VAR_GLOBAL CONSTANT   // PLC tag table "Open Library"
   "Modes.Auto" : Int := 1;
   "Modes.Manual" : Int := 2;
   "Modes.Independent" : Int := 10;
   "Modes.Stop" : Int := 0;
   "HMI.Status.Stopped" : Int := 0;
   "HMI.Status.Estop" : Int := 1;
   "HMI.Status.Error" : Int := 2;
   "HMI.Status.ForwardWork" : Int := 3;
   "HMI.Status.ReverseHome" : Int := 4;
   "HMI.Status.OnForwardWork" : Int := 5;
   "HMI.Status.OnReverseHome" : Int := 6;
   "IoScaling.S7Analog.Default.iRawMax" : Int := 27648;
   "IoScaling.S7Analog.Default.iRawMin" : Int := 0;
   "IoScaling.S7Analog.Default.bSwapBytes" : Bool := false;
   "IoScaling.S7Analog.+-V/mA.iRawMax" : Int := 27648;
   "IoScaling.S7Analog.+-V/mA.iRawMin" : Int := -27648;
   "IoScaling.S7Analog.Types.Default" : Int := 0;
   "IoScaling.S7Analog.Pt100.iRawMax" : Int := 8500;
   "IoScaling.S7Analog.Pt100.iRawMin" : Int := -2000;
   "IoScaling.S7Analog.Pt100.Climate.iRawMax" : Int := 13000;
   "IoScaling.S7Analog.Pt100.Climate.iRawMin" : Int := -12000;
   "IoScaling.S7Analog.Ni100.iRawMax" : Int := 2500;
   "IoScaling.S7Analog.Ni100.iRawMin" : Int := -600;
   "IoScaling.S7Analog.Ni100.Climate.iRawMax" : Int := 25000;
   "IoScaling.S7Analog.Ni100.Climate.iRawMin" : Int := -6000;
   "IoScaling.S7Analog.Types.+-V/mA" : Int := 1;
   "IoScaling.S7Analog.Types.Pt100" : Int := 2;
   "IoScaling.S7Analog.Types.Pt100.Climate" : Int := 3;
   "IoScaling.S7Analog.Types.Ni100" : Int := 4;
   "IoScaling.S7Analog.Types.Ni100.Climate" : Int := 5;
   "IoScaling.S7Analog.Pt100.rScaledMax" : Real := 850.0;
   "IoScaling.S7Analog.Pt100.rScaledMin" : Real := -200.0;
   "IoScaling.S7Analog.Pt100.Climate.rScaledMax" : Real := 130.0;
   "IoScaling.S7Analog.Pt100.Climate.rScaledMin" : Real := -120.0;
   "IoScaling.S7Analog.Ni100.rScaledMax" : Real := 250.0;
   "IoScaling.S7Analog.Ni100.rScaledMin" : Real := -60.0;
   "IoScaling.S7Analog.Ni100.Climate.rScaledMax" : Real := 250.0;
   "IoScaling.S7Analog.Ni100.Climate.rScaledMin" : Real := -60.0;
   "IoScaling.S7Analog.150Ohms.rScaledMax" : Real := 150.0;
   "IoScaling.S7Analog.150Ohms.rScaledMin" : Real := 0.0;
   "IoScaling.S7Analog.300Ohms.rScaledMax" : Real := 300.0;
   "IoScaling.S7Analog.300Ohms.rScaledMin" : Real := 0.0;
   "IoScaling.S7Analog.600Ohms.rScaledMax" : Real := 600.0;
   "IoScaling.S7Analog.600Ohms.rScaledMin" : Real := 0.0;
   "Estop.MinSetPoint" : Int := 0;
   "Estop.MaxSetPoint" : Int := 1;
   "Estop.HMISetPoint" : Int := 2;
   "Modes.PID.Inactive" : Int := 0;
   "Modes.PID.Pretuning" : Int := 1;
   "Modes.PID.FineTuning" : Int := 2;
   "Modes.PID.AutoMode" : Int := 3;
   "Modes.PID.ManualMode" : Int := 4;
   "HMI.Status.Generic1" : Int := 101;
   "HMI.Status.Generic2" : Int := 102;
   "HMI.Status.Generic3" : Int := 103;
   "HMI.Status.Generic4" : Int := 104;
   "HMI.Status.Generic5" : Int := 105;
   "HMI.Status.GenericNone" : Int := 100;
   "HMI.Status.Generic6" : Int := 106;
   "DataTypes.rMaxReal" : Real := 3.402823e38;
   "DataTypes.rMinReal" : Real := -3.402823e38;
   "DataTypes.iMaxInt" : Int := 32767;
   "DataTypes.iMinInt" : Int := -32768;
END_VAR

(* ===== HMI "HMI_RT_1" =====
connection "HMI_Connection_1": ETHERNET, S7_1500_OMS

HMI tags "Default tag table"
   "Tag_ScreenNumber" : UInt, internal
   "dbErrors_WaterSystem" : Array [0..49] of Word, 1 s
   "dbWaterSystem_AI_WaterPumpPressure" : udtHMI_AnalogInput, 1 s
   "dbWaterSystem_WaterTemperature_AI_WaterTemperature" : udtHMI_AnalogInput, 1 s
   "dbWaterSystem_MTR_ReturnWaterPump" : udtHMI_MotorControl, 1 s
   "dbWaterSystem_ANA_SteamValve" : udtHMI_AnalogValveControl, 1 s
   "dbWaterSystem_VFD_WaterPump" : udtHMI_VFD_Control, 1 s
   "dbWaterSystem_SOL_MainWater" : udtHMI_ValveControl, 1 s
   "dbWaterSystem_AO_CoolingCoil" : udtHMI_AnalogOutput, 1 s
   "dbWaterSystem_AO_CoolingCoil_rValue" : Real, 1 s
   "dbErrors_AirSystem" : Array [0..1] of Word, 1 s
   "dbWaterSystem_SystemControl" : udtHMI_SystemControl, 1 s
   "dbAirSystem_VFD_RecirculationFan" : udtHMI_VFD_Control, 1 s
   "dbAirSystem_SystemControl" : udtHMI_SystemControl, 1 s

HMI tags "PID"
   "dbWaterSystem_WaterTemperature_PID_WaterTempInterface" : udtHMI_PIDInterface, 1 s

discrete alarms
   1: '', class Errors, trigger "dbErrors_WaterSystem" bit 8
   2: '', class Errors, trigger "dbErrors_WaterSystem" bit 9
   3: '', class Errors, trigger "dbErrors_WaterSystem" bit 10
   4: '', class Errors, trigger "dbErrors_WaterSystem" bit 11
   5: '', class Errors, trigger "dbErrors_WaterSystem" bit 24
   6: '', class Errors, trigger "dbErrors_WaterSystem" bit 25
   7: '', class Errors, trigger "dbErrors_WaterSystem" bit 26
   8: '', class Errors, trigger "dbErrors_WaterSystem" bit 27
   9: '', class Errors, trigger "dbErrors_WaterSystem" bit 28
   10: '', class Errors, trigger "dbErrors_WaterSystem" bit 29
   11: '', class Errors, trigger "dbErrors_WaterSystem" bit 30
   12: '', class Errors, trigger "dbErrors_WaterSystem" bit 31
   13: '', class Errors, trigger "dbErrors_WaterSystem" bit 16
   14: '', class Errors, trigger "dbErrors_WaterSystem" bit 17
   15: '', class Errors, trigger "dbErrors_WaterSystem" bit 18
   16: '', class Errors, trigger "dbErrors_WaterSystem" bit 19
   17: '', class Errors, trigger "dbErrors_WaterSystem" bit 20
   18: '', class Errors, trigger "dbErrors_WaterSystem" bit 21
   19: '', class Errors, trigger "dbErrors_WaterSystem" bit 40
   20: '', class Errors, trigger "dbErrors_WaterSystem" bit 41
   21: '', class Errors, trigger "dbErrors_WaterSystem" bit 42
   22: '', class Errors, trigger "dbErrors_WaterSystem" bit 56
   23: '', class Errors, trigger "dbErrors_WaterSystem" bit 57
   24: '', class Errors, trigger "dbErrors_WaterSystem" bit 58
   25: '', class Errors, trigger "dbErrors_WaterSystem" bit 59
   26: '', class Errors, trigger "dbErrors_WaterSystem" bit 60
   27: '', class Errors, trigger "dbErrors_WaterSystem" bit 61
   28: '', class Errors, trigger "dbErrors_WaterSystem" bit 72
   29: '', class Errors, trigger "dbErrors_WaterSystem" bit 88
   30: '', class Errors, trigger "dbErrors_WaterSystem" bit 89
   31: '', class Errors, trigger "dbErrors_WaterSystem" bit 104
   32: '', class Errors, trigger "dbErrors_WaterSystem" bit 105
   33: '', class Errors, trigger "dbErrors_WaterSystem" bit 106
   34: '', class Errors, trigger "dbErrors_WaterSystem" bit 107
   35: '', class Errors, trigger "dbErrors_WaterSystem" bit 108
   36: '', class Errors, trigger "dbErrors_WaterSystem" bit 109
   37: '', class Errors, trigger "dbErrors_WaterSystem" bit 110
   38: '', class Errors, trigger "dbErrors_WaterSystem" bit 111
   39: '', class Errors, trigger "dbErrors_WaterSystem" bit 96
   40: '', class Errors, trigger "dbErrors_WaterSystem" bit 97
   41: '', class Errors, trigger "dbErrors_WaterSystem" bit 98
   42: '', class Errors, trigger "dbErrors_WaterSystem" bit 99
   43: '', class Errors, trigger "dbErrors_WaterSystem" bit 100
   44: '', class Errors, trigger "dbErrors_WaterSystem" bit 101
   45: '', class Errors, trigger "dbErrors_WaterSystem" bit 102
   46: '', class Errors, trigger "dbErrors_WaterSystem" bit 120
   47: '', class Errors, trigger "dbErrors_WaterSystem" bit 121
   48: '', class Errors, trigger "dbErrors_WaterSystem" bit 122
   49: '', class Errors, trigger "dbErrors_WaterSystem" bit 136
   50: '', class Errors, trigger "dbErrors_WaterSystem" bit 137
   51: '', class Errors, trigger "dbErrors_AirSystem" bit 8
   52: '', class Errors, trigger "dbErrors_AirSystem" bit 9
   53: '', class Errors, trigger "dbErrors_AirSystem" bit 10
   54: '', class Errors, trigger "dbErrors_AirSystem" bit 11
   55: '', class Errors, trigger "dbErrors_AirSystem" bit 12
   56: '', class Errors, trigger "dbErrors_AirSystem" bit 13
   57: '', class Errors, trigger "dbErrors_AirSystem" bit 14
   58: '', class Errors, trigger "dbErrors_AirSystem" bit 15
   59: '', class Errors, trigger "dbErrors_AirSystem" bit 0
   60: '', class Errors, trigger "dbErrors_AirSystem" bit 1
   61: '', class Errors, trigger "dbErrors_AirSystem" bit 2
   62: '', class Errors, trigger "dbErrors_AirSystem" bit 3
   63: '', class Errors, trigger "dbErrors_AirSystem" bit 4
   64: '', class Errors, trigger "dbErrors_AirSystem" bit 5

screen "Water System" 800x480, template "Template"
   SymbolLibrary "Symbol library_18" at 288,346 size 39x53
   SymbolLibrary "Symbol library_16" at 609,374 size 40x40
   SymbolLibrary "Symbol library_15" at 590,249 size 40x40
   SymbolLibrary "Symbol library_13" at 446,334 size 58x20
   SymbolLibrary "Symbol library_12" at 341,238 size 44x9
   SymbolLibrary "Symbol library_11" at 437,238 size 44x9
   SymbolLibrary "Symbol library_10" at 533,249 size 63x21
   SymbolLibrary "Symbol library_8" at 246,334 size 128x20
   SymbolLibrary "Symbol library_4" at 73,264 size 21x72
   SymbolLibrary "Symbol library_2" at 74,115 size 40x40
   SymbolLibrary "Symbol library_1" at 25,148 size 118x198
   TextField "Text field_1" at 42,201 size 83x42
   SymbolLibrary "Symbol library_3" at 73,334 size 40x40
   SymbolLibrary "Symbol library_5" at 106,354 size 55x20
   SymbolLibrary "Symbol library_6" at 111,115 size 344x21
   SymbolLibrary "Symbol library_7" at 535,95 size 98x21
   ScreenModuleView "fpMotor_Pump_Horizontal_1" at 440,79 size 109x91
   TextField "Text field_2" at 646,117 size 66x38
   ScreenModuleView "fpVFD_Pump_Horizontal_1" at 149,317 size 109x92
   SymbolLibrary "Symbol library_9" at 478,230 size 64x155
   TextField "Text field_3" at 407,398 size 98x21
   ScreenModuleView "fpValve_Analog_Horizontal_1" at 369,178 size 80x87
   TextField "Text field_4" at 265,254 size 54x21
   ScreenModuleView "fpValve_Solenoid_Horizontal_1" at 356,311 size 93x68
   SymbolLibrary "Symbol library_14" at 592,281 size 68x102
   TextField "Text field_5" at 675,237 size 58x38
   Bar "Bar_1" at 599,286 size 40x92
   SymbolLibrary "Symbol library_17" at 642,394 size 55x20
   TextField "Text field_6" at 714,350 size 65x38
   Button "Button_1" at 439,79 size 110x91
   Button "Button_2" at 149,317 size 110x91
   Button "Button_3" at 369,178 size 80x87
   Button "Button_4" at 356,311 size 93x68
   Button "Button_5" at 591,279 size 71x104
   ScreenModuleView "fp_AnalogInput_Numeric_1" at 265,408 size 88x31
   SymbolLibrary "Symbol library_19" at 565,214 size 38x35
   ScreenModuleView "fp_AnalogInput_Numeric_2" at 533,178 size 88x31
   ScreenModuleView "fp_AnalogOutput_1" at 663,295 size 70x41
   ScreenModuleView "fpModeControl_1" at 0,0 size 170x70
   Button "Button_6" at 260,347 size 95x94
   Button "Button_7" at 530,174 size 95x86
   Button "Button_8" at 0,0 size 170x70
   Button "Button_9" at 698,1 size 102x70

Template "Template" 800x480
   Button "Template_Button" at 720,422 size 78x58
   AlarmView "Alarm view_1" at 170,1 size 529x70

PopupScreen "AI Main Water Pump Pressure" 220x253
   ScreenModuleView "fpIO_AnalogInput_Popup_1" at 0,0 size 220x253
   Button "Button_5" at 115,217 size 95x26

PopupScreen "MTR Return Water Pump" 180x300
   ScreenModuleView "fpMotor_Reversing_Popup_1" at 0,0 size 180x300
   Button "Button_5" at 95,264 size 75x26

PopupScreen "SOL Main Water Valve" 180x272
   ScreenModuleView "fpValve_Solenoid_Popup_1" at 0,0 size 180x272
   Button "Button_5" at 97,236 size 71x26

PopupScreen "ANA Water Temperature Valve" 220x277
   ScreenModuleView "fpValve_Analog_Popup_1" at 0,0 size 220x277
   Button "Button_5" at 113,241 size 95x26

PopupScreen "VFD Main Water Pump" 180x387
   ScreenModuleView "fpVFD_Popup" at 0,0 size 180x387
   Button "Button_5" at 98,350 size 71x26

PopupScreen "AO Cooling Coil" 220x275
   ScreenModuleView "fpIO_AnalogOutput_Popup_1" at 0,0 size 220x275
   Button "Button_5" at 114,236 size 95x26

PopupScreen "SYS Water System" 180x285
   ScreenModuleView "fpModeControl_Popup_1" at 0,0 size 180x285
   Button "Button_5" at 99,249 size 71x26

PopupScreen "AI Main Water Temperature" 220x253
   ScreenModuleView "fpIO_AnalogInput_Popup_1" at 0,0 size 220x253
   Button "Button_5" at 115,217 size 95x26

screen "Air System" 800x480, template "Template"
   ScreenModuleView "fpModeControl_1" at 0,0 size 170x70
   Button "Button_8" at 0,0 size 170x70
   Button "Button_9" at 698,1 size 102x70
   SymbolLibrary "Symbol library_6" at 343,83 size 185x61
   SymbolLibrary "Symbol library_2" at 223,83 size 122x120
   SymbolLibrary "Symbol library_3" at 223,335 size 122x120
   TextField "Text field_2" at 546,107 size 64x38
   TextField "Text field_6" at 551,389 size 63x38
   SymbolLibrary "Symbol library_1" at 343,394 size 185x61
   SymbolLibrary "Symbol library_4" at 223,299 size 62x37
   SymbolLibrary "Symbol library_5" at 224,202 size 62x37
   GraphicView "Graphic view_1" at 224,238 size 61x61
   ScreenModuleView "fpVFD_Motor_Horizontal_1" at 90,230 size 139x77
   Button "Button_2" at 90,230 size 139x77

PopupScreen "SYS Air System" 180x285
   ScreenModuleView "fpModeControl_Popup_1" at 0,0 size 180x285
   Button "Button_5" at 99,249 size 71x26

PopupScreen "VFD Air Recirculation Fan" 180x387
   ScreenModuleView "fpAir_Recirculation_VFD_Popup" at 0,0 size 180x387
   Button "Button_5" at 98,350 size 71x26
*)

(* ===== HMI "HMI_RT_1" =====

ScreenModuleEditorView "fpInterlock" 640x480
   GraphicView "Graphic view_1" at 231,83 size 200x200
*)

(* ===== HMI "HMI_RT_1" =====

text list "ErrorMessages": 0..1 ''; 1 ''; 2 ''; 3 ''

text list "InterlockList": 0 ''; 1 ''

text list "InterlockIndicators": 0 ''; 1 ''; 2 ''

ScreenModuleEditorView "fpInterlock8_Popup" 640x480
   TextField "Text field_1" at 10,12 size 180x31
   IOField "I/O field_1" at 20,47 size 150x20
   IOField "I/O field_2" at 20,67 size 150x20
   IOField "I/O field_3" at 20,87 size 150x20
   IOField "I/O field_4" at 20,107 size 150x20
   IOField "I/O field_5" at 20,127 size 150x20
   IOField "I/O field_6" at 20,147 size 150x20
   IOField "I/O field_7" at 20,167 size 150x20
   IOField "I/O field_8" at 20,187 size 150x20
   SymbolicIOField "Symbolic I/O field_3" at 126,47 size 54x20
   SymbolicIOField "Symbolic I/O field_1" at 126,67 size 54x20
   SymbolicIOField "Symbolic I/O field_2" at 126,87 size 54x20
   SymbolicIOField "Symbolic I/O field_4" at 126,107 size 54x20
   SymbolicIOField "Symbolic I/O field_5" at 126,127 size 54x20
   SymbolicIOField "Symbolic I/O field_6" at 126,147 size 54x20
   SymbolicIOField "Symbolic I/O field_7" at 126,167 size 54x20
   SymbolicIOField "Symbolic I/O field_8" at 126,187 size 54x20
*)

(* ===== HMI "HMI_RT_1" =====

text list "ErrorMessages": 0..1 ''; 1 ''; 2 ''; 3 ''

text list "InterlockList": 0 ''; 1 ''

text list "InterlockIndicators": 0 ''; 1 ''; 2 ''

ScreenModuleEditorView "fpInterlock16_Popup" 640x480
   TextField "Text field_1" at 10,12 size 180x31
   IOField "I/O field_1" at 20,47 size 150x20
   IOField "I/O field_2" at 20,67 size 150x20
   IOField "I/O field_3" at 20,87 size 150x20
   IOField "I/O field_4" at 20,107 size 150x20
   IOField "I/O field_5" at 20,127 size 150x20
   IOField "I/O field_6" at 20,147 size 150x20
   IOField "I/O field_7" at 20,167 size 150x20
   IOField "I/O field_8" at 20,187 size 150x20
   IOField "I/O field_9" at 20,207 size 150x20
   IOField "I/O field_10" at 20,227 size 150x20
   IOField "I/O field_11" at 20,247 size 150x20
   IOField "I/O field_12" at 20,267 size 150x20
   IOField "I/O field_13" at 20,287 size 150x20
   IOField "I/O field_14" at 20,307 size 150x20
   IOField "I/O field_15" at 20,327 size 150x20
   IOField "I/O field_16" at 20,347 size 150x20
   SymbolicIOField "Symbolic I/O field_3" at 126,47 size 54x20
   SymbolicIOField "Symbolic I/O field_1" at 126,67 size 54x20
   SymbolicIOField "Symbolic I/O field_2" at 126,87 size 54x20
   SymbolicIOField "Symbolic I/O field_4" at 126,107 size 54x20
   SymbolicIOField "Symbolic I/O field_5" at 126,127 size 54x20
   SymbolicIOField "Symbolic I/O field_6" at 126,147 size 54x20
   SymbolicIOField "Symbolic I/O field_7" at 126,167 size 54x20
   SymbolicIOField "Symbolic I/O field_8" at 126,187 size 54x20
   SymbolicIOField "Symbolic I/O field_9" at 126,207 size 54x20
   SymbolicIOField "Symbolic I/O field_10" at 126,227 size 54x20
   SymbolicIOField "Symbolic I/O field_11" at 126,247 size 54x20
   SymbolicIOField "Symbolic I/O field_12" at 126,267 size 54x20
   SymbolicIOField "Symbolic I/O field_13" at 126,287 size 54x20
   SymbolicIOField "Symbolic I/O field_14" at 126,307 size 54x20
   SymbolicIOField "Symbolic I/O field_15" at 126,327 size 54x20
   SymbolicIOField "Symbolic I/O field_16" at 126,347 size 54x20
*)

(* ===== HMI "HMI_RT_1" =====

text list "ErrorMessages": 0 ''; 1 ''

text list "IndependantMode": 0 ''; 1 ''

text list "EStop": 0 ''; 1 ''

text list "Auto": 0 ''; 1 ''

ScreenModuleEditorView "fpSystemControl_Popup" 640x480
   Button "Button_1" at 20,50 size 159x28
   Button "Button_4" at 20,261 size 71x26
   Button "Button_2" at 20,87 size 160x28
   SymbolicIOField "Symbolic I/O field_3" at 20,195 size 160x25
   TextField "Text field_1" at 10,12 size 180x31
   SymbolicIOField "Symbolic I/O field_5" at 20,228 size 160x25
   Button "Button_3" at 20,122 size 160x28
   Button "Button_6" at 20,158 size 160x28
*)

(* ===== HMI "HMI_RT_1" =====

text list "ErrorMessages": 0..1 ''; 1 ''; 2 ''; 3 ''

text list "InterlockList": 0 ''; 1 ''

text list "InterlockIndicators": 0 ''; 1 ''; 2 ''

ScreenModuleEditorView "fpInterlock8_Popup_s7_300" 640x480
   TextField "Text field_1" at 10,12 size 180x31
   IOField "I/O field_1" at 20,47 size 150x20
   IOField "I/O field_2" at 20,67 size 150x20
   IOField "I/O field_3" at 20,87 size 150x20
   IOField "I/O field_4" at 20,107 size 150x20
   IOField "I/O field_5" at 20,127 size 150x20
   IOField "I/O field_6" at 20,147 size 150x20
   IOField "I/O field_7" at 20,167 size 150x20
   IOField "I/O field_8" at 20,187 size 150x20
   SymbolicIOField "Symbolic I/O field_3" at 126,47 size 54x20
   SymbolicIOField "Symbolic I/O field_1" at 126,67 size 54x20
   SymbolicIOField "Symbolic I/O field_2" at 126,87 size 54x20
   SymbolicIOField "Symbolic I/O field_4" at 126,107 size 54x20
   SymbolicIOField "Symbolic I/O field_5" at 126,127 size 54x20
   SymbolicIOField "Symbolic I/O field_6" at 126,147 size 54x20
   SymbolicIOField "Symbolic I/O field_7" at 126,167 size 54x20
   SymbolicIOField "Symbolic I/O field_8" at 126,187 size 54x20
*)

(* ===== HMI "HMI_RT_1" =====

text list "ErrorMessages": 0..1 ''; 1 ''; 2 ''; 3 ''

text list "InterlockList": 0 ''; 1 ''

text list "InterlockIndicators": 0 ''; 1 ''; 2 ''

ScreenModuleEditorView "fpInterlock16_Popup_s7_300" 640x480
   TextField "Text field_1" at 10,12 size 180x31
   IOField "I/O field_1" at 20,47 size 150x20
   IOField "I/O field_2" at 20,67 size 150x20
   IOField "I/O field_3" at 20,87 size 150x20
   IOField "I/O field_4" at 20,107 size 150x20
   IOField "I/O field_5" at 20,127 size 150x20
   IOField "I/O field_6" at 20,147 size 150x20
   IOField "I/O field_7" at 20,167 size 150x20
   IOField "I/O field_8" at 20,187 size 150x20
   IOField "I/O field_9" at 20,207 size 150x20
   IOField "I/O field_10" at 20,227 size 150x20
   IOField "I/O field_11" at 20,247 size 150x20
   IOField "I/O field_12" at 20,267 size 150x20
   IOField "I/O field_13" at 20,287 size 150x20
   IOField "I/O field_14" at 20,307 size 150x20
   IOField "I/O field_15" at 20,327 size 150x20
   IOField "I/O field_16" at 20,347 size 150x20
   SymbolicIOField "Symbolic I/O field_3" at 126,47 size 54x20
   SymbolicIOField "Symbolic I/O field_1" at 126,67 size 54x20
   SymbolicIOField "Symbolic I/O field_2" at 126,87 size 54x20
   SymbolicIOField "Symbolic I/O field_4" at 126,107 size 54x20
   SymbolicIOField "Symbolic I/O field_5" at 126,127 size 54x20
   SymbolicIOField "Symbolic I/O field_6" at 126,147 size 54x20
   SymbolicIOField "Symbolic I/O field_7" at 126,167 size 54x20
   SymbolicIOField "Symbolic I/O field_8" at 126,187 size 54x20
   SymbolicIOField "Symbolic I/O field_9" at 126,207 size 54x20
   SymbolicIOField "Symbolic I/O field_10" at 126,227 size 54x20
   SymbolicIOField "Symbolic I/O field_11" at 126,247 size 54x20
   SymbolicIOField "Symbolic I/O field_12" at 126,267 size 54x20
   SymbolicIOField "Symbolic I/O field_13" at 126,287 size 54x20
   SymbolicIOField "Symbolic I/O field_14" at 126,307 size 54x20
   SymbolicIOField "Symbolic I/O field_15" at 126,327 size 54x20
   SymbolicIOField "Symbolic I/O field_16" at 126,347 size 54x20
*)

(* ===== HMI "HMI_RT_1" =====

text list "InterlockList": 0 ''; 1 ''

text list "ErrorMessages": 0..1 ''; 5 ''; 6 ''; 7 ''; 8 ''; 9 ''; 10 ''; 11 ''; 12 ''; 13 ''; 14 ''; 15 ''; 16 ''; 17 ''; 18 ''; 19 ''

ScreenModuleEditorView "fpPID_CompactInterace_Popup_s7_300" 640x480
   Button "Button_1" at 20,50 size 95x28
   Button "Button_4" at 20,351 size 95x26
   TextField "Text field_4" at 20,86 size 23x15
   IOField "I/O field_1" at 43,84 size 72x18
   TextField "Text field_5" at 125,86 size 23x15
   IOField "I/O field_2" at 147,84 size 72x18
   TextField "Text field_6" at 20,135 size 66x15
   TextField "Text field_7" at 20,113 size 59x15
   IOField "I/O field_3" at 120,112 size 100x17
   IOField "I/O field_4" at 120,134 size 100x17
   Button "Button_2" at 125,50 size 95x28
   SymbolicIOField "Symbolic I/O field_3" at 19,316 size 200x24
   TextField "Text field_1" at 10,12 size 220x31
   TextField "Text field_2" at 20,157 size 60x15
   IOField "I/O field_6" at 120,156 size 100x17
   TextField "Text field_8" at 20,214 size 14x15
   IOField "I/O field_7" at 34,212 size 81x18
   TextField "Text field_9" at 20,236 size 12x15
   IOField "I/O field_8" at 34,234 size 81x18
   TextField "Text field_10" at 20,258 size 15x15
   IOField "I/O field_9" at 34,256 size 81x18
   TextField "Text field_11" at 125,214 size 22x15
   IOField "I/O field_10" at 147,212 size 73x18
   TextField "Text field_12" at 125,236 size 23x15
   IOField "I/O field_11" at 147,234 size 73x18
   Button "Button_3" at 20,280 size 60x26
   Button "Button_6" at 90,280 size 60x26
   Button "Button_7" at 160,280 size 60x26
   Button "Button_8" at 20,183 size 95x24
   Button "Button_9" at 125,183 size 95x24
*)

(* ===== HMI "HMI_RT_1" =====

text list "InterlockList": 0 ''; 1 ''

text list "ErrorMessages": 0..1 ''; 5 ''; 6 ''; 7 ''; 8 ''; 9 ''; 10 ''; 11 ''; 12 ''; 13 ''; 14 ''; 15 ''; 16 ''; 17 ''; 18 ''; 19 ''

ScreenModuleEditorView "fpPID_CompactInterface_Popup_Graph_s7_300" 640x480
   Button "Button_1" at 20,50 size 95x28
   Button "Button_4" at 20,426 size 95x26
   TextField "Text field_4" at 20,86 size 23x15
   IOField "I/O field_1" at 43,84 size 72x18
   TextField "Text field_5" at 125,86 size 23x15
   IOField "I/O field_2" at 147,84 size 72x18
   TextField "Text field_6" at 20,137 size 66x15
   TextField "Text field_7" at 20,116 size 59x15
   IOField "I/O field_3" at 120,115 size 100x17
   IOField "I/O field_4" at 120,136 size 100x17
   Button "Button_2" at 125,50 size 95x28
   SymbolicIOField "Symbolic I/O field_3" at 20,188 size 420x24
   TextField "Text field_1" at 10,12 size 440x30
   TextField "Text field_2" at 20,157 size 60x15
   IOField "I/O field_6" at 120,157 size 100x17
   TextField "Text field_8" at 238,86 size 14x15
   IOField "I/O field_7" at 252,84 size 81x18
   TextField "Text field_9" at 238,108 size 12x15
   IOField "I/O field_8" at 252,106 size 81x18
   TextField "Text field_10" at 238,130 size 15x15
   IOField "I/O field_9" at 252,128 size 81x18
   TextField "Text field_11" at 343,86 size 22x15
   IOField "I/O field_10" at 365,84 size 73x18
   TextField "Text field_12" at 343,108 size 23x15
   IOField "I/O field_11" at 365,106 size 73x18
   Button "Button_3" at 238,152 size 60x26
   Button "Button_6" at 308,152 size 60x26
   Button "Button_7" at 378,152 size 60x26
   Button "Button_8" at 238,50 size 95x28
   Button "Button_9" at 343,50 size 95x28
   TrendView "Trend view_1" at 20,226 size 420x195
*)

(* ===== HMI "HMI_RT_1" =====

text list "ErrorMessages": 0 ''; 1 ''

text list "IndependantMode": 0 ''; 1 ''

text list "EStop": 0 ''; 1 ''

text list "Auto": 0 ''; 1 ''

ScreenModuleEditorView "fpSystemControl_Popup_s7_300" 640x480
   Button "Button_1" at 20,50 size 159x28
   Button "Button_4" at 20,261 size 71x26
   Button "Button_2" at 20,87 size 160x28
   SymbolicIOField "Symbolic I/O field_3" at 20,195 size 160x25
   TextField "Text field_1" at 10,12 size 180x31
   SymbolicIOField "Symbolic I/O field_5" at 20,228 size 160x25
   Button "Button_3" at 20,122 size 160x28
   Button "Button_6" at 20,158 size 160x28
*)

(* ===== HMI "HMI_RT_1" =====

ScreenModuleEditorView "fp_AnalogInput_Numeric_s7_300" 640x480
   IOField "I/O field_1" at 27,18 size 100x25
*)

(* ===== HMI "HMI_RT_1" =====

ScreenModuleEditorView "fp_AnalogOutput_s7_300" 640x480
   IOField "I/O field_1" at 159,73 size 96x32
   GraphicView "Graphic view_1" at 190,73 size 34x32
*)

(* ===== HMI "HMI_RT_1" =====

ScreenModuleEditorView "fpMotor_Motor_Horizontal_s7_300" 640x480
   SymbolLibrary "Symbol library_3" at 167,75 size 165x85
   GraphicView "Graphic view_1" at 204,77 size 80x80
*)

(* ===== HMI "HMI_RT_1" =====

ScreenModuleEditorView "fpMotor_Motor_Vertical_s7_300" 640x480
   SymbolLibrary "Symbol library_3" at 59,35 size 85x165
   GraphicView "Graphic view_1" at 61,83 size 80x80
*)

(* ===== HMI "HMI_RT_1" =====

ScreenModuleEditorView "fpMotor_Pump_Horizontal_s7_300" 640x480
   SymbolLibrary "Symbol library_3" at 208,75 size 125x85
   GraphicView "Graphic view_1" at 231,84 size 70x70
*)

(* ===== HMI "HMI_RT_1" =====

ScreenModuleEditorView "fpMotor_Pump_Vertical_s7_300" 640x480
   SymbolLibrary "Symbol library_3" at 19,24 size 85x125
   GraphicView "Graphic view_1" at 28,56 size 70x70
*)

(* ===== HMI "HMI_RT_1" =====

ScreenModuleEditorView "fpValve_Analog_Horizontal_s7_300" 640x480
   SymbolLibrary "Symbol library_1" at 34,25 size 165x165
   Bar "Bar_1" at 57,84 size 119x38
   GraphicView "Graphic view_1" at 81,120 size 70x70
*)

(* ===== HMI "HMI_RT_1" =====

ScreenModuleEditorView "fpValve_Analog_Vertical_s7_300" 640x480
   SymbolLibrary "Symbol library_1" at 39,27 size 165x165
   Bar "Bar_1" at 99,55 size 40x110
   GraphicView "Graphic view_1" at 132,74 size 70x70
*)

(* ===== HMI "HMI_RT_1" =====

ScreenModuleEditorView "fpValve_Solenoid_Horizontal_s7_300" 640x480
   SymbolLibrary "Symbol library_1" at 21,17 size 165x85
   GraphicView "Graphic view_1" at 69,24 size 70x70
*)

(* ===== HMI "HMI_RT_1" =====

ScreenModuleEditorView "fpValve_Solenoid_Vertical_s7_300" 640x480
   SymbolLibrary "Symbol library_1" at 16,18 size 85x165
   GraphicView "Graphic view_1" at 24,66 size 70x70
*)

(* ===== HMI "HMI_RT_1" =====

ScreenModuleEditorView "fpVFD_Motor_Horizontal_s7_300" 640x480
   SymbolLibrary "Symbol library_3" at 167,75 size 165x85
   GraphicView "Graphic view_1" at 210,78 size 80x80
*)

(* ===== HMI "HMI_RT_1" =====

ScreenModuleEditorView "fpVFD_Motor_Vertical_s7_300" 640x480
   SymbolLibrary "Symbol library_3" at 59,35 size 85x165
   GraphicView "Graphic view_1" at 62,78 size 80x80
*)

(* ===== HMI "HMI_RT_1" =====

ScreenModuleEditorView "fpVFD_Pump_Horizontal_s7_300" 640x480
   SymbolLibrary "Symbol library_3" at 208,75 size 125x85
   GraphicView "Graphic view_1" at 231,83 size 70x70
*)

(* ===== HMI "HMI_RT_1" =====

ScreenModuleEditorView "fpVFD_Pump_Vertical_s7_300" 640x480
   SymbolLibrary "Symbol library_3" at 19,24 size 85x125
   GraphicView "Graphic view_1" at 27,55 size 70x70
*)

(* ===== HMI "HMI_RT_1" =====

ScreenModuleEditorView "fpInterlock_s7_300" 640x480
   GraphicView "Graphic view_1" at 231,83 size 200x200
*)

(* ===== HMI "HMI_RT_1" =====

text list "SystemModes": 1 ''; 2 ''; 10 ''; 0 ''

ScreenModuleEditorView "fpSystemControl_s7_300" 640x480
   TextField "Text field_1" at 85,10 size 170x70
   SymbolicIOField "Symbolic I/O field_1" at 95,40 size 150x30
*)

(* ===== HMI "HMI_RT_1" =====

text list "HMIStatus": 0..1 ''; 101 ''; 102 ''; 103 ''; 104 ''; 105 ''

text list "InterlockList": 0 ''; 1 ''

ScreenModuleEditorView "fpIO_AnalogInput_Popup_s7_300" 640x480
   Button "Button_1" at 20,50 size 95x28
   Button "Button_4" at 20,229 size 95x26
   TextField "Text field_4" at 20,130 size 57x15
   IOField "I/O field_1" at 110,128 size 110x20
   TextField "Text field_5" at 32,93 size 72x15
   IOField "I/O field_2" at 135,90 size 75x20
   Button "Button_2" at 125,50 size 95x28
   SymbolicIOField "Symbolic I/O field_3" at 20,189 size 200x24
   TextField "Text field_1" at 10,12 size 220x31
   TextField "Text field_2" at 20,158 size 62x15
   IOField "I/O field_3" at 110,157 size 110x20
*)

(* ===== HMI "HMI_RT_1" =====

text list "ErrorMessages": 0..1 ''; 1 ''; 2 ''; 3 ''

text list "InterlockList": 0 ''; 1 ''

ScreenModuleEditorView "fpIO_AnalogOutput_Popup_s7_300" 640x480
   Button "Button_1" at 20,50 size 95x28
   Button "Button_4" at 20,248 size 95x26
   TextField "Text field_5" at 125,89 size 23x15
   IOField "I/O field_2" at 147,88 size 72x18
   Button "Button_2" at 125,50 size 95x28
   SymbolicIOField "Symbolic I/O field_1" at 20,176 size 200x24
   SymbolicIOField "Symbolic I/O field_3" at 19,208 size 200x24
   TextField "Text field_1" at 10,12 size 220x31
   TextField "Text field_7" at 21,123 size 60x15
   IOField "I/O field_1" at 120,122 size 100x18
   TextField "Text field_2" at 20,89 size 23x15
   IOField "I/O field_3" at 42,88 size 72x18
   TextField "Text field_3" at 21,147 size 61x15
   IOField "I/O field_4" at 120,146 size 100x18
*)

(* ===== HMI "HMI_RT_1" =====

text list "InterlockList": 1 ''; 0 ''; 2 ''

text list "ErrorMessages": 0..1 ''; 1 ''; 2 ''; 3 ''; 4 ''; 5 ''; 6 ''; 7 ''

ScreenModuleEditorView "fpMotor_Reversing_Popup_s7_300" 640x480
   Button "Button_1" at 20,50 size 75x28
   Button "Button_3" at 26,172 size 148x27
   Button "Button_4" at 20,276 size 75x26
   Button "Button_6" at 26,203 size 148x28
   Button "Button_7" at 26,235 size 148x28
   Button "Button_2" at 105,50 size 75x28
   SymbolicIOField "Symbolic I/O field_1" at 20,94 size 160x24
   SymbolicIOField "Symbolic I/O field_3" at 20,126 size 160x24
   TextField "Text field_1" at 10,12 size 180x31
*)

(* ===== HMI "HMI_RT_1" =====

text list "InterlockList": 1 ''; 0 ''

text list "ErrorMessages": 0..1 ''; 1 ''; 2 ''

ScreenModuleEditorView "fpValve_Analog_Popup_s7_300" 640x480
   SymbolicIOField "Symbolic I/O field_1" at 19,183 size 200x24
   Button "Button_1" at 20,50 size 95x28
   Button "Button_4" at 20,253 size 95x26
   TextField "Text field_4" at 20,88 size 23x15
   IOField "I/O field_1" at 43,86 size 72x18
   TextField "Text field_5" at 125,88 size 23x15
   IOField "I/O field_2" at 147,86 size 72x18
   TextField "Text field_7" at 20,146 size 34x15
   IOField "I/O field_3" at 120,145 size 100x17
   Button "Button_2" at 125,50 size 95x28
   SymbolicIOField "Symbolic I/O field_3" at 19,212 size 200x24
   TextField "Text field_1" at 10,12 size 220x31
   TextField "Text field_2" at 20,113 size 48x15
   IOField "I/O field_4" at 120,112 size 100x17
*)

(* ===== HMI "HMI_RT_1" =====

text list "InterlockList": 1 ''; 0 ''; 2 ''

text list "ErrorMessages": 0..1 ''; 1 ''; 2 ''; 3 ''; 5 ''; 4 ''

ScreenModuleEditorView "fpValve_Solenoid_Popup_s7_300" 640x480
   Button "Button_1" at 20,50 size 75x28
   Button "Button_4" at 20,248 size 71x26
   Button "Button_2" at 104,50 size 75x28
   SymbolicIOField "Symbolic I/O field_1" at 20,94 size 159x24
   SymbolicIOField "Symbolic I/O field_3" at 19,126 size 159x24
   TextField "Text field_1" at 10,12 size 180x31
   Button "Button_8" at 24,174 size 148x27
   Button "Button_9" at 23,205 size 148x27
*)

(* ===== HMI "HMI_RT_1" =====

text list "InterlockList": 1 ''; 0 ''

text list "ErrorMessages": 4 ''; 1 ''; 2 ''; 3 ''; 5 ''; 6 ''; 7 ''; 8 ''; 9 ''; 10 ''; 11 ''; 12 ''; 13 ''; 14 ''; 15 ''; 15 ''

ScreenModuleEditorView "fpVFD_Popup_s7_300" 640x480
   Button "Button_1" at 20,50 size 75x28
   Button "Button_3" at 25,258 size 148x27
   Button "Button_4" at 20,362 size 71x26
   Button "Button_6" at 25,288 size 148x28
   Button "Button_7" at 25,320 size 148x28
   TextField "Text field_4" at 16,92 size 23x15
   IOField "I/O field_1" at 39,90 size 56x18
   TextField "Text field_5" at 99,92 size 23x15
   IOField "I/O field_2" at 121,90 size 57x18
   TextField "Text field_6" at 21,152 size 68x15
   TextField "Text field_7" at 21,130 size 63x15
   IOField "I/O field_3" at 88,129 size 91x17
   IOField "I/O field_4" at 88,151 size 91x17
   Button "Button_2" at 104,50 size 75x28
   SymbolicIOField "Symbolic I/O field_1" at 20,182 size 159x24
   SymbolicIOField "Symbolic I/O field_3" at 19,213 size 159x24
   TextField "Text field_1" at 10,12 size 180x31
*)

(* ===== HMI "HMI_RT_1" =====

ScreenModuleEditorView "fp_AnalogInput_Numeric" 640x480
   IOField "I/O field_1" at 27,18 size 100x25
*)

(* ===== HMI "HMI_RT_1" =====

ScreenModuleEditorView "fp_AnalogOutput" 640x480
   IOField "I/O field_1" at 159,73 size 96x32
   GraphicView "Graphic view_1" at 190,73 size 34x32
*)

(* ===== HMI "HMI_RT_1" =====

ScreenModuleEditorView "fpMotor_Motor_Vertical" 640x480
   SymbolLibrary "Symbol library_3" at 59,35 size 85x165
   GraphicView "Graphic view_1" at 61,83 size 80x80
*)

(* ===== HMI "HMI_RT_1" =====

ScreenModuleEditorView "fpMotor_Pump_Horizontal" 640x480
   SymbolLibrary "Symbol library_3" at 208,75 size 125x85
   GraphicView "Graphic view_1" at 231,84 size 70x70
*)

(* ===== HMI "HMI_RT_1" =====

ScreenModuleEditorView "fpMotor_Pump_Vertical" 640x480
   SymbolLibrary "Symbol library_3" at 19,24 size 85x125
   GraphicView "Graphic view_1" at 28,56 size 70x70
*)

(* ===== HMI "HMI_RT_1" =====

ScreenModuleEditorView "fpMotor_Motor_Horizontal" 640x480
   SymbolLibrary "Symbol library_3" at 167,75 size 165x85
   GraphicView "Graphic view_1" at 204,77 size 80x80
*)

(* ===== HMI "HMI_RT_1" =====

ScreenModuleEditorView "fpValve_Analog_Vertical" 640x480
   SymbolLibrary "Symbol library_1" at 39,27 size 165x165
   Bar "Bar_1" at 99,55 size 40x110
   GraphicView "Graphic view_1" at 132,74 size 70x70
*)

(* ===== HMI "HMI_RT_1" =====

ScreenModuleEditorView "fpValve_Analog_Horizontal" 640x480
   SymbolLibrary "Symbol library_1" at 34,25 size 165x165
   Bar "Bar_1" at 57,84 size 119x38
   GraphicView "Graphic view_1" at 81,120 size 70x70
*)

(* ===== HMI "HMI_RT_1" =====

ScreenModuleEditorView "fpValve_Solenoid_Horizontal" 640x480
   SymbolLibrary "Symbol library_1" at 21,17 size 165x85
   GraphicView "Graphic view_1" at 69,24 size 70x70
*)

(* ===== HMI "HMI_RT_1" =====

ScreenModuleEditorView "fpValve_Solenoid_Vertical" 640x480
   SymbolLibrary "Symbol library_1" at 16,18 size 85x165
   GraphicView "Graphic view_1" at 24,66 size 70x70
*)

(* ===== HMI "HMI_RT_1" =====

ScreenModuleEditorView "fpVFD_Motor_Horizontal" 640x480
   SymbolLibrary "Symbol library_3" at 167,75 size 165x85
   GraphicView "Graphic view_1" at 210,78 size 80x80
*)

(* ===== HMI "HMI_RT_1" =====

ScreenModuleEditorView "fpVFD_Motor_Vertical" 640x480
   SymbolLibrary "Symbol library_3" at 59,35 size 85x165
   GraphicView "Graphic view_1" at 62,78 size 80x80
*)

(* ===== HMI "HMI_RT_1" =====

ScreenModuleEditorView "fpVFD_Pump_Horizontal" 640x480
   SymbolLibrary "Symbol library_3" at 208,75 size 125x85
   GraphicView "Graphic view_1" at 231,83 size 70x70
*)

(* ===== HMI "HMI_RT_1" =====

ScreenModuleEditorView "fpVFD_Pump_Vertical" 640x480
   SymbolLibrary "Symbol library_3" at 19,24 size 85x125
   GraphicView "Graphic view_1" at 27,55 size 70x70
*)

(* ===== HMI "HMI_RT_1" =====

text list "SystemModes": 1 ''; 2 ''; 10 ''; 0 ''

ScreenModuleEditorView "fpSystemControl" 640x480
   TextField "Text field_1" at 85,10 size 170x70
   SymbolicIOField "Symbolic I/O field_1" at 95,40 size 150x30
*)

(* ===== HMI "HMI_RT_1" =====

text list "HMIStatus": 0..1 ''; 101 ''; 102 ''; 103 ''; 104 ''; 105 ''

text list "InterlockList": 0 ''; 1 ''

ScreenModuleEditorView "fpIO_AnalogInput_Popup" 640x480
   Button "Button_1" at 20,50 size 95x28
   Button "Button_4" at 20,229 size 95x26
   TextField "Text field_4" at 20,130 size 57x15
   IOField "I/O field_1" at 110,128 size 110x20
   TextField "Text field_5" at 32,93 size 72x15
   IOField "I/O field_2" at 135,90 size 75x20
   Button "Button_2" at 125,50 size 95x28
   SymbolicIOField "Symbolic I/O field_3" at 20,189 size 200x24
   TextField "Text field_1" at 10,12 size 220x31
   TextField "Text field_2" at 20,158 size 62x15
   IOField "I/O field_3" at 110,157 size 110x20
*)

(* ===== HMI "HMI_RT_1" =====

text list "ErrorMessages": 0..1 ''; 1 ''; 2 ''; 3 ''

text list "InterlockList": 0 ''; 1 ''

ScreenModuleEditorView "fpIO_AnalogOutput_Popup" 640x480
   Button "Button_1" at 20,50 size 95x28
   Button "Button_4" at 20,248 size 95x26
   TextField "Text field_5" at 125,89 size 23x15
   IOField "I/O field_2" at 147,88 size 72x18
   Button "Button_2" at 125,50 size 95x28
   SymbolicIOField "Symbolic I/O field_1" at 20,176 size 200x24
   SymbolicIOField "Symbolic I/O field_3" at 19,208 size 200x24
   TextField "Text field_1" at 10,12 size 220x31
   TextField "Text field_7" at 21,123 size 60x15
   IOField "I/O field_1" at 120,122 size 100x18
   TextField "Text field_2" at 20,89 size 23x15
   IOField "I/O field_3" at 42,88 size 72x18
   TextField "Text field_3" at 21,147 size 61x15
   IOField "I/O field_4" at 120,146 size 100x18
*)

(* ===== HMI "HMI_RT_1" =====

text list "InterlockList": 1 ''; 0 ''; 2 ''

text list "ErrorMessages": 0..1 ''; 1 ''; 2 ''; 3 ''; 4 ''; 5 ''; 6 ''; 7 ''

ScreenModuleEditorView "fpMotor_Reversing_Popup" 640x480
   Button "Button_1" at 20,50 size 75x28
   Button "Button_3" at 26,172 size 148x27
   Button "Button_4" at 20,276 size 75x26
   Button "Button_6" at 26,203 size 148x28
   Button "Button_7" at 26,235 size 148x28
   Button "Button_2" at 105,50 size 75x28
   SymbolicIOField "Symbolic I/O field_1" at 20,94 size 160x24
   SymbolicIOField "Symbolic I/O field_3" at 20,126 size 160x24
   TextField "Text field_1" at 10,12 size 180x31
*)

(* ===== HMI "HMI_RT_1" =====

text list "InterlockList": 0 ''; 1 ''

text list "ErrorMessages": 0..1 ''; 1 ''; 2 ''

ScreenModuleEditorView "fpValve_Analog_Popup" 640x480
   SymbolicIOField "Symbolic I/O field_1" at 19,183 size 200x24
   Button "Button_1" at 20,50 size 95x28
   Button "Button_4" at 20,253 size 95x26
   TextField "Text field_4" at 20,88 size 23x15
   IOField "I/O field_1" at 43,86 size 72x18
   TextField "Text field_5" at 125,88 size 23x15
   IOField "I/O field_2" at 147,86 size 72x18
   TextField "Text field_7" at 20,146 size 34x15
   IOField "I/O field_3" at 120,145 size 100x17
   Button "Button_2" at 125,50 size 95x28
   SymbolicIOField "Symbolic I/O field_3" at 19,212 size 200x24
   TextField "Text field_1" at 10,12 size 220x31
   TextField "Text field_2" at 20,113 size 48x15
   IOField "I/O field_4" at 120,112 size 100x17
*)

(* ===== HMI "HMI_RT_1" =====

text list "InterlockList": 1 ''; 0 ''; 2 ''

text list "ErrorMessages": 0..1 ''; 1 ''; 2 ''; 3 ''; 4 ''; 5 ''

ScreenModuleEditorView "fpValve_Solenoid_Popup" 640x480
   Button "Button_1" at 20,50 size 75x28
   Button "Button_4" at 20,248 size 71x26
   Button "Button_2" at 104,50 size 75x28
   SymbolicIOField "Symbolic I/O field_1" at 21,94 size 159x24
   SymbolicIOField "Symbolic I/O field_3" at 21,126 size 159x24
   TextField "Text field_1" at 10,12 size 180x31
   Button "Button_8" at 26,174 size 148x27
   Button "Button_9" at 26,205 size 148x27
*)

(* ===== HMI "HMI_RT_1" =====

text list "InterlockList": 1 ''; 0 ''

text list "ErrorMessages": 0..1 ''; 1 ''; 2 ''; 3 ''; 4 ''; 5 ''; 6 ''; 7 ''; 8 ''; 9 ''; 10 ''; 11 ''; 12 ''; 13 ''; 14 ''; 15 ''

ScreenModuleEditorView "fpVFD_Popup" 640x480
   Button "Button_1" at 20,50 size 75x28
   Button "Button_3" at 25,258 size 148x27
   Button "Button_4" at 20,362 size 71x26
   Button "Button_6" at 25,288 size 148x28
   Button "Button_7" at 25,320 size 148x28
   TextField "Text field_4" at 16,92 size 23x15
   IOField "I/O field_1" at 39,90 size 56x18
   TextField "Text field_5" at 99,92 size 23x15
   IOField "I/O field_2" at 121,90 size 57x18
   TextField "Text field_6" at 21,152 size 68x15
   TextField "Text field_7" at 21,130 size 63x15
   IOField "I/O field_3" at 88,129 size 91x17
   IOField "I/O field_4" at 88,151 size 91x17
   Button "Button_2" at 104,50 size 75x28
   SymbolicIOField "Symbolic I/O field_1" at 20,182 size 159x24
   SymbolicIOField "Symbolic I/O field_3" at 19,213 size 159x24
   TextField "Text field_1" at 10,12 size 180x31
*)

(* ===== HMI "HMI_RT_1" =====

text list "InterlockList": 0 ''; 1 ''

text list "ErrorMessages": 0..1 ''; 1 ''; 2 ''; 3 ''; 4 ''; 5 ''; 6 ''; 7 ''; 8 ''; 9 ''; 10 ''; 11 ''; 12 ''; 13 ''; 14 ''; 15 ''; 16 ''

ScreenModuleEditorView "fpPID_CompactInterface_Popup_Graph" 640x480
   Button "Button_1" at 20,50 size 95x28
   Button "Button_4" at 20,426 size 95x26
   TextField "Text field_4" at 20,86 size 23x15
   IOField "I/O field_1" at 43,84 size 72x18
   TextField "Text field_5" at 125,86 size 23x15
   IOField "I/O field_2" at 147,84 size 72x18
   TextField "Text field_6" at 20,138 size 66x15
   TextField "Text field_7" at 20,116 size 59x15
   IOField "I/O field_3" at 120,115 size 100x17
   IOField "I/O field_4" at 120,137 size 100x17
   Button "Button_2" at 125,50 size 95x28
   SymbolicIOField "Symbolic I/O field_3" at 20,188 size 420x24
   TextField "Text field_1" at 10,12 size 440x30
   TextField "Text field_2" at 20,160 size 60x15
   IOField "I/O field_6" at 120,159 size 100x17
   TextField "Text field_8" at 238,86 size 14x15
   IOField "I/O field_7" at 252,84 size 81x18
   TextField "Text field_9" at 238,108 size 12x15
   IOField "I/O field_8" at 252,106 size 81x18
   TextField "Text field_10" at 238,130 size 15x15
   IOField "I/O field_9" at 252,128 size 81x18
   TextField "Text field_11" at 343,86 size 22x15
   IOField "I/O field_10" at 365,84 size 73x18
   TextField "Text field_12" at 343,108 size 23x15
   IOField "I/O field_11" at 365,106 size 73x18
   Button "Button_3" at 238,152 size 60x26
   Button "Button_6" at 308,152 size 60x26
   Button "Button_7" at 378,152 size 60x26
   Button "Button_8" at 238,50 size 95x28
   Button "Button_9" at 343,50 size 95x28
   TrendView "Trend view_1" at 20,230 size 420x195
*)

(* ===== HMI "HMI_RT_1" =====

text list "InterlockList": 0 ''; 1 ''

text list "ErrorMessages": 0..1 ''; 1 ''; 2 ''; 3 ''; 4 ''; 5 ''; 6 ''; 7 ''; 8 ''; 9 ''; 10 ''; 11 ''; 12 ''; 13 ''; 14 ''; 15 ''; 16 ''

ScreenModuleEditorView "fpPID_CompactInterace_Popup" 640x480
   Button "Button_1" at 20,50 size 95x28
   Button "Button_4" at 20,349 size 95x26
   TextField "Text field_4" at 20,86 size 23x15
   IOField "I/O field_1" at 43,84 size 72x18
   TextField "Text field_5" at 125,86 size 23x15
   IOField "I/O field_2" at 147,84 size 72x18
   TextField "Text field_6" at 20,134 size 66x15
   TextField "Text field_7" at 20,113 size 59x15
   IOField "I/O field_3" at 120,112 size 100x17
   IOField "I/O field_4" at 120,133 size 100x17
   Button "Button_2" at 125,50 size 95x28
   SymbolicIOField "Symbolic I/O field_3" at 19,314 size 200x24
   TextField "Text field_1" at 10,12 size 220x31
   TextField "Text field_2" at 20,156 size 60x15
   IOField "I/O field_6" at 120,155 size 100x17
   TextField "Text field_8" at 20,212 size 14x15
   IOField "I/O field_7" at 34,210 size 81x18
   TextField "Text field_9" at 20,234 size 12x15
   IOField "I/O field_8" at 34,232 size 81x18
   TextField "Text field_10" at 20,256 size 15x15
   IOField "I/O field_9" at 34,254 size 81x18
   TextField "Text field_11" at 125,212 size 22x15
   IOField "I/O field_10" at 147,210 size 73x18
   TextField "Text field_12" at 125,234 size 23x15
   IOField "I/O field_11" at 147,232 size 73x18
   Button "Button_3" at 20,278 size 60x26
   Button "Button_6" at 90,278 size 60x26
   Button "Button_7" at 160,278 size 60x26
   Button "Button_8" at 20,181 size 95x24
   Button "Button_9" at 125,181 size 95x24
*)